
   ResetOfNotifyROS:R     "Notity_for_Rotor_over_speed";
         JU    Brake_Failure;


   //BRAKE FAILURE ALARM
   Brake_Failure:A     "Alarm_reset";
         FP    #os11;
         JC    ResetOfAlaramBF;
         CLR;
         A     "Notify_reset";
         FP    #os12;
         JC    ResetOfNotifyBF;
         CLR;
         L     "rotor_rpm";
         L     0;
         >I;
         L     "Brake_Out_HOA";
         JC    TIMERFORBF;
         JU    E_STOP;
   TIMERFORBF:CALL  "Convert_time"
         ( iv1   := "BrakeFailureSP",
           time1 := #TI_6
         );
         CALL  TON , "IEC_Timer_0_DB_24"
         ( IN := true,
           PT := #TI_6,
           Q  := #BF_AT,
           ET := #T6
         );
         A     #BF_AT;
         JC    SetOfAlarmBF;
         JU    E_STOP;

   SetOfAlarmBF:SET;
         S     "Alarm_for_Brake_failure";
         S     "Notity_for_Brake_failure";
         JU    E_STOP;
   ResetOfAlaramBF:R     "Alarm_for_Brake_failure";
         R     "Notity_for_Brake_failure";
         CALL  RESET_TIMER
         ( "TIMER" := "IEC_Timer_0_DB_24"
         );
         JU    E_STOP;
   ResetOfNotifyBF:R     "Notity_for_Brake_failure";
         JU    E_STOP;


   // E_STOP ALARM
   E_STOP:A     "Alarm_reset";
         FP    #os14;
         JC    ResetOfAlaramES;
         CLR;
         A     "Notify_reset";
         FP    #os15;
         JC    ResetOfNotifyES;
         CLR;
         A     "E_Stop";
         JC    SetOfAlarmES;
         JU    AlarmCtrl;

   SetOfAlarmES:SET;
         S     "Alarm_for_E_Stop";
         S     "Notity_for_E_Stop";
         JU    AlarmCtrl;

   ResetOfAlaramES:R     "Alarm_for_E_Stop";
         R     "Notity_for_E_Stop";
         JU    AlarmCtrl;
   ResetOfNotifyES:R     "Notity_for_E_Stop";
         JU    AlarmCtrl;

   // Alarm Horn Ctrl
   AlarmCtrl:A     "Fault_Mode";
         FP    #os16;
         JC    AlarmCtrl_SET;
         CLR;
         A     "Alarm_reset";
         O     "Notify_reset";
         FP    #os17;
         JC    ResetAlarmCtrl;
         JU    End_of_line;

   AlarmCtrl_SET:SET;
         S     "Alarm_CTRL";
         JU    End_of_line;

   ResetAlarmCtrl:R     "Alarm_CTRL";
         JU    End_of_line;

   End_of_line:BE;
END_REGION
END_FUNCTION_BLOCK

FUNCTION_BLOCK "Modes_STL"   // FB17, STL
{ S7_Optimized_Access := 'TRUE' }
VERSION : 0.1
   VAR
      os1 : Bool;
      os2 : Bool;
   END_VAR
   VAR_TEMP
      ti1 : Time;
      WarmUpTrigger : Bool;
      tm1 : Time;
      tv1 : Int;
      tv2 : Int;
      tb1 : Bool;
      ti2 : Time;
      Stabilizetrigger : Bool;
      tm2 : Time;
      ti3 : Time;
      CooldownTrigger : Bool;
      tm3 : Time;
   END_VAR
BEGIN

REGION Network 1
   // ESTOP HANDLING
         A     "Alarm_for_E_Stop";
         O     "Alarm_for_Brake_failure";
         JC    EstopAlarm;
         JU    Reset_EStopAlarm;

   EstopAlarm:SET;
         S     "Warm_Transition";
         S     "Stabilize_Transition";
         S     "Generation_Transition";
         S     "CoolDown_Transition";

   Reset_EStopAlarm:CLR;
         R     "Warm_Transition";
         R     "Stabilize_Transition";
         R     "Generation_Transition";
         R     "CoolDown_Transition";

   JumpToMode:A     "Warm_UP_Mode";
         JC    Start_WarmUp;
         CLR;
         A     "Stabilize_mode";
         JC    StabilizeMode;
         CLR;
         A     "Generation_Mode";
         JC    GenerationMode;
         CLR;
         A     "CoolDown_Mode";
         JC    CooldownMode;
         CLR;
         A     "Idle_Mode";
         JC    IdleMode;
         JU    EndOfLine;


   // WARM UP MODE
   Start_WarmUp:SET;
         R     "Warm_Transition";
         R     "Stabilize_Transition";
         R     "Generation_Transition";
         R     "CoolDown_Transition";
         R     "StartSequenceBit";
         CLR;
         A     "Warm_UP_Mode";
         JC    WarmUpMode;
         CLR;
         A     "Stabilize_mode";
         JC    StabilizeMode;
         CLR;
         A     "Generation_Mode";
         JC    GenerationMode;
         CLR;
         A     "CoolDown_Mode";
         JC    CooldownMode;
         CLR;
         A     "Idle_Mode";
         JC    IdleMode;
         JU    EndOfLine;

   WarmUpMode:SET;
         NOT;
         R     "Brake_Out_CTRL";
         L     "Warmup_RPM";
         T     "BafflePID_SP";
         L     "rotor_rpm";
         T     "BafflePIDin";

         SET;
         S     "OilPumpVFD_CTRL";
         S     "Baffle_Ctrl";
         L     "WarmUp_VFDper";
         T     "VFDsp";

         L     "Oil_temp";
         L     "WarmUpOilTempSp";
         >I;
         JC    WarmUpMode;
         CALL  RESET_TIMER
         ( "TIMER" := "IEC_Timer_0_DB_35"
         );
         JU    StabilizeMode;

   WarmUpTime:CALL  "Convert_time"
         ( iv1   := "WarmUpOilDelaySp",
           time1 := #ti1
         );
         CALL  TON, "IEC_Timer_0_DB_35"
         ( IN := true,
           PT := #ti1,
           Q  := #WarmUpTrigger,
           ET := #tm1
         );
         A     #WarmUpTrigger;
         JC    WarmUpExit;
         CLR;
         A     "Alarm_for_Rotor_over_speed";
         O     "Alarm_for_High_temp";
         JC    WarmUpExit;
         JU    StabilizeMode;

   WarmUpExit:S     "Warm_Transition";
         CALL  RESET_TIMER
         ( "TIMER" := "IEC_Timer_0_DB_35"
         );
         JU    StabilizeMode;


   //STABILZE MODE
   StabilizeMode:SET;
         NOT;
         R     "Warm_Transition";
         L     "StabilizekWSP";
         T     "BafflePID_SP";
         L     "Current_flow";
         T     "BafflePIDin";
         L     "StabilizekWSP";
         L     5;
         +I;
         T     #tv1;
         T     "StabilizekWSP";
         L     5;
         -I;
         L     #tv2;
         L     "Current_flow";
         L     #tv1;
         <I;
         S     #tb1;
         L     "Current_flow";
         L     #tv2;
         >I;
         A     #tb1;
         JC    StabilizeMode;
         CALL  RESET_TIMER
         ( "TIMER" := "IEC_Timer_0_DB_36"
         );
         JU    GenerationMode;
   StabilizeTime:CALL  "Convert_time"
         ( iv1   := "StabilizeDealySP",
           time1 := #ti2
         );
         CALL  TON, "IEC_Timer_0_DB_36"
         ( IN := true,
           PT := #ti2,
           Q  := #Stabilizetrigger,
           ET := #tm2
         );
         A     #Stabilizetrigger;
         JC    StabilizeExit;
         CLR;
         A     "Alarm_for_Rotor_over_speed";
         O     "Alarm_for_High_temp";
         JC    StabilizeExit;
         JU    GenerationMode;

   StabilizeExit:S     "Stabilize_Transition";
         CALL  RESET_TIMER
         ( "TIMER" := "IEC_Timer_0_DB_36"
         );
         JU    GenerationMode;


   //GENERATION MODE
   GenerationMode:SET;
         NOT;
         R     "Stabilize_Transition";
         SET;
         S     "Station_Interlock_CTRL";
         A     "System_Stop_PB";
         JC    GenerationExit;
         CLR;
         A     "Alarm_for_Over_Current";
         JC    GenerationExit;
         CLR;
         A     "Alarm_for_Rotor_over_speed";
         O     "Alarm_for_High_temp";
         JC    GenerationExit;
         JU    CooldownMode;

   GenerationExit:S     "Generation_Transition";
         JU    CooldownMode;


   //COOLDOWN MODE
   CooldownMode:SET;
         NOT;
         R     "Generation_Transition";
         R     "Station_Interlock_CTRL";
         L     "CoolDown_RPM";
         T     "BafflePID_SP";
         L     "rotor_rpm";
         T     "BafflePIDin";
         L     "Oil_temp";
         L     "CoolDownOilTempSp";
         <I;
         JC    Cooldowntime;
         CALL  RESET_TIMER
         ( "TIMER" := "IEC_Timer_0_DB_37"
         );
         JU    IdleMode;

   Cooldowntime:CALL  "Convert_time"
         ( iv1   := "CoolDownlDelaySp",
           time1 := #ti3
         );
         CALL  TON, "IEC_Timer_0_DB_37"
         ( IN := true,
           PT := #ti3,
           Q  := #CooldownTrigger,
           ET := #tm3
         );
         A     #CooldownTrigger;
         JC    CooldownExit;
         JU    IdleMode;

   CooldownExit:S     "CoolDown_Transition";
         CALL  RESET_TIMER
         ( "TIMER" := "IEC_Timer_0_DB_37"
         );
         JU    IdleMode;


   //IDLE MODE
   IdleMode:SET;
         NOT;
         R     "CoolDown_Transition";
         R     "Station_Interlock_CTRL";
         S     "Brake_Out_CTRL";
         R     "Baffle_Ctrl";
         R     "OilPumpVFD_CTRL";
         CLR;
         A     "StartSequencePB";
         A     "Idle_Mode";
         A     "FULLAUTOBIT";
         FP    #os2;
         S     "StartSequenceBit";
         JU    EndOfLine;

   //FAULT MODE
   EndOfLine:A     "E_Stop";
         O     "Alarm_for_Brake_failure";
         O     "Alarm_for_High_temp";
         O     "Alarm_for_LOW_OIL";
         O     "Alarm_for_Oil_High_Flow";
         O     "Alarm_for_Over_Current";
         O     "Alarm_for_Rotor_over_speed";
         =     "Fault_Mode";
END_REGION
END_FUNCTION_BLOCK

FUNCTION_BLOCK "HOURMETER_STL"   // FB22, STL
{ S7_Optimized_Access := 'TRUE' }
VERSION : 0.1
   VAR
      Min_time_down : Bool;
      Min_countdown : Bool;
      Hour_countdown : Bool;
      Day_countdown : Bool;
      Day_count_down : Bool;
      Hr_count_down : Bool;
      reset_rto : Bool;
      min_count_reset : Bool;
      hour_count_reset : Bool;
      reset_hourmeter_trigger : Bool;
      os3 : Bool;
      os2 : Bool;
      os1 : Bool;
      os4 : Bool;
      Reset_HM_Trigger : Bool;
      accum_elapsed : Time;
   END_VAR
   VAR_TEMP
      resettime : Time;
      toooomanydays : Bool;
   END_VAR
BEGIN

REGION Network 1
         A     "Generation_Mode";
         JC    RTOtimer;
         CLR;
         A     "Reset_HM_PB";
         JC    RestHourmeter;
         JU    EndOfLine;

   RTOtimer:CALL  TONR , "IEC_Timer_0_DB_44"
         ( IN := true,
           R  := #reset_rto,
           PT := t#1m,
           Q  := #Min_time_down,
           ET := #accum_elapsed
         );

         CALL  CTU, "n"
         ( CU := #Min_countdown,
           R  := #min_count_reset,
           PV := 60,
           Q  := #Hr_count_down,
           CV := "HM_Minutes"
         );

         CALL  CTU, "IEC_Counter_0_DB_9"
         ( CU := #Hour_countdown,
           R  := #hour_count_reset,
           PV := 24,
           Q  := #Day_count_down,
           CV := "HM_Hours"
         );

         CALL  CTU, "nt"
         ( CU := #Day_countdown,
           R  := #reset_hourmeter_trigger,
           PV := 10000,
           Q  := #toooomanydays,
           CV := "HM_Days"
         );

         JU    EndOfLine;

   RestHourmeter:CALL  TON, "IEC_Timer_0_DB_45"
         ( IN := "Reset_HM_PB",
           PT := T#10s,
           Q  := #Reset_HM_Trigger,
           ET := #resettime
         );

   EndOfLine:CLR;
         A     #Reset_HM_Trigger;
         O     #Min_countdown;
         =     #reset_rto;
         CLR;
         A     #Reset_HM_Trigger;
         O     #Hour_countdown;
         =     #min_count_reset;
         CLR;
         A     #Reset_HM_Trigger;
         O     #Day_countdown;
         =     #hour_count_reset;
         CLR;
END_REGION
END_FUNCTION_BLOCK

(* ===== HMI "HMI_RT_1" =====
system functions are stored by id; their names below are inferred from use
connection "1500": ETHERNET, S7_1500_OMS

HMI tags "Default tag table"
   "StartSequencePB" : Bool = PLC StartSequencePB AT %M43.7, 1 s
   "System_Stop_PB" : Bool = PLC System_Stop_PB AT %M48.7, 1 s
   "Alarm_for_E_Stop" : Bool = PLC Alarm_for_E_Stop AT %M56.0, 1 s
   "Alarm_for_Brake_failure" : Bool = PLC Alarm_for_Brake_failure AT %M55.7, 1 s
   "Alarm_for_High_temp" : Bool = PLC Alarm_for_High_temp AT %M29.7, 1 s
   "Alarm_for_LOW_OIL" : Bool = PLC Alarm_for_LOW_OIL AT %M30.0, 1 s
   "Alarm_for_Oil_High_Flow" : Bool = PLC Alarm_for_Oil_High_Flow AT %M30.1, 1 s
   "Alarm_for_Over_Current" : Bool = PLC Alarm_for_Over_Current AT %M30.2, 1 s
   "Alarm_for_Rotor_over_speed" : Bool = PLC Alarm_for_Rotor_over_speed AT %M30.3, 1 s
   "Alarm_HAND_PB" : Bool = PLC Alarm_HAND_PB AT %M28.5, 1 s
   "Alarm_HOA" : Int = PLC Alarm_HOA AT %MW34, 1 s
   "Alarm_OFF_PB" : Bool = PLC Alarm_OFF_PB AT %M28.4, 1 s
   "Alarm_reset" : Bool = PLC Alarm_reset AT %M29.6, 1 s
   "Baffle_Out" : Int = PLC Baffle_Out AT %MW18, 1 s
   "Baffle_AUTO_PB" : Bool = PLC Baffle_AUTO_PB AT %M81.2, 1 s
   "Baffle_HAND_PB" : Bool = PLC Baffle_HAND_PB AT %M81.0, 1 s
   "Baffle_HOA" : Int = PLC Baffle_HOA AT %MW94, 1 s
   "Baffle_Manual" : Bool = PLC Baffle_Manual AT %M96.0, 1 s
   "Baffle_OFF_PB" : Bool = PLC Baffle_OFF_PB AT %M81.1, 1 s
   "Brake_AUTO_PB" : Bool = PLC Brake_AUTO_PB AT %M28.3, 1 s
   "Brake_HAND_PB" : Bool = PLC Brake_HAND_PB AT %M28.2, 1 s
   "Brake_OFF_PB" : Bool = PLC Brake_OFF_PB AT %M28.1, 1 s
   "Brake_Out" : Bool = PLC Brake_Out AT %M0.0, 1 s
   "Brake_Out_CTRL" : Bool = PLC Brake_Out_CTRL AT %M29.3, 1 s
   "Brake_Out_HOA" : Int = PLC Brake_Out_HOA AT %MW32, 1 s
   "Station_interlock_HAND_PB" : Bool = PLC Station_interlock_HAND_PB AT %M29.0, 1 s
   "Station_Interlock_HOA" : Int = PLC Station_Interlock_HOA AT %MW36, 1 s
   "Station_interlock_OFF_PB" : Bool = PLC Station_interlock_OFF_PB AT %M28.7, 1 s
   "Station_interlock_AUTO_PB" : Bool = PLC Station_interlock_AUTO_PB AT %M29.1, 1 s
   "Station_interlock" : Bool = PLC Station_interlock AT %M1.3, 1 s
   "VFD_HOA" : Int = PLC VFD_HOA AT %MW98, 1 s
   "VFDHOA_AUTO_PB" : Bool = PLC VFDHOA_AUTO_PB AT %M96.1, 1 s
   "VFDHOA_HAND_PB" : Bool = PLC VFDHOA_HAND_PB AT %M96.3, 1 s
   "VFDHOA_OFF_PB" : Bool = PLC VFDHOA_OFF_PB AT %M96.2, 1 s
   "Notify_reset" : Bool = PLC Notify_reset AT %M42.1, 1 s
   "Fault_Mode" : Bool = PLC Fault_Mode AT %M80.4, 1 s
   "HighOilTempDelaySP" : Int = PLC HighOilTempDelaySP AT %MW64, 1 s
   "HM_Days" : Int = PLC HM_Days AT %MW108, 1 s
   "HM_Hours" : Int = PLC HM_Hours AT %MW106, 1 s
   "HM_Minutes" : Int = PLC HM_Minutes AT %MW30, 1 s
   "ModeInt" : Int = PLC ModeInt AT %MW110, 1 s
   "OverCurrenDelaytSP" : Int = PLC OverCurrenDelaytSP AT %MW44, 1 s
   "OilHighFlowSP" : Int = PLC OilHighFlowSP AT %MW58, 1 s
   "OilLowFlowDelaySP" : Int = PLC OilLowFlowDelaySP AT %MW38, 1 s
   "RotorOverSpeedSP" : Int = PLC RotorOverSpeedSP AT %MW54, 1 s
   "WarmUpOilTemp" : Int = PLC WarmUpOilTempSp AT %MW74, 1 s
   "CoolDownlDelaySp" : Int = PLC CoolDownlDelaySp AT %MW84, 1 s
   "CoolDownOilTemp" : Int = PLC CoolDownOilTempSp AT %MW86, 1 s
   "StabilizeDealySP" : Int = PLC StabilizeDealySP AT %MW78, 1 s
   "Alarm_horn_Q" : Bool = PLC Alarm_horn_Q AT %M1.4, 1 s
   "ManualBaffle_SP" : Real = PLC ManualBaffle_SP AT %MD90, 1 s
   "ManualVFD_SP" : Real = PLC ManualVFD_SP AT %MD100, 1 s
   "Alarm_HighOilTemp_int" : Int = PLC Alarm_HighOilTemp_int AT %MW112, 1 s
   "Alarm_LowOilFlow_int" : Int = PLC Alarm_LowOilFlow_int AT %MW114, 1 s
   "Alarm_HighOilFlow_int" : Int = PLC Alarm_HighOilFlow_int AT %MW116, 1 s
   "Alarm_OverCurrent_int" : Int = PLC Alarm_OverCurrent_int AT %MW118, 1 s
   "Alarm_RotorOverSpeed_int" : Int = PLC Alarm_RotorOverSpeed_int AT %MW120, 1 s
   "Alarm_BrakeFailure_int" : Int = PLC Alarm_BrakeFailure_int AT %MW122, 1 s
   "Alarm_EStop_int" : Int = PLC Alarm_EStop_int AT %MW124, 1 s
   "ProgramLanguage" : Int = PLC Program_lang AT %MW12, 1 s
   "LADpb" : Bool = PLC PB_LAD AT %M0.4, 1 s
   "FBDpb" : Bool = PLC PB_FBD AT %M0.5, 1 s
   "SCLpb" : Bool = PLC PB_SCL AT %M0.6, 1 s
   "STLpb" : Bool = PLC PB_STL AT %M0.7, 1 s
   "Current" : Int = PLC Current_flow AT %MW26, 1 s
   "Oil Flow" : Int = PLC Oil_flow AT %MW22, 1 s
   "Oil temp" : Int = PLC Oil_temp AT %MW24, 1 s
   "BrakeFailuredelay" : Int = PLC BrakeFailureSP AT %MW60, 1 s
   "Rpm sp" : Int = PLC Rotor_Over_SpeedSp AT %MW56, 1 s
   "OverSpeedSP" : Int = PLC RotorOverSpeedSP AT %MW54, 1 s
   "Warmup delay" : Int = PLC WarmUpOilDelaySp AT %MW72, 1 s
   "AlarmAuto_Pb" : Bool = PLC Alarm_AUTO_PB AT %M28.6, 1 s
   "RPM" : Int = PLC rotor_rpm AT %MW20, 1 s
   "OilPct" : Int = PLC Oil_pump_vfd_per AT %MW14, 1 s
   "baffle" : Int = PLC Baffle_per AT %MW16, 1 s
   "brakeEN" : Bool = PLC Brake_Out AT %M0.0, 1 s
   "InterlockEN" : Bool = PLC Station_interlock AT %M1.3, 1 s
   "HM reset" : Bool = PLC Reset_HM_PB AT %M49.0, 1 s
   "currentdealy" : Int = PLC OverCurrenDelaytSP AT %MW44, 1 s
   "high oil temp sp" : Int = PLC High_Oil_TempSp AT %MW52, 1 s
   "low oil flow sp" : Int = PLC Oil_lowSp AT %MW40, 1 s
   "curent sp" : Int = PLC Over_currentSp AT %MW46, 1 s
   "high oil flow sp" : Int = PLC Oil_highSp AT %MW62, 1 s

discrete alarms
   1: 'EStop Activated', class Errors, trigger "Alarm_EStop_int" bit 0
   2: 'Low Oil Flow Alert', class Errors, trigger "Alarm_LowOilFlow_int" bit 0
   3: 'Over Current Alert', class Errors, trigger "Alarm_OverCurrent_int" bit 0
   4: 'High Oil Temperature Alert', class Errors, trigger "Alarm_HighOilTemp_int" bit 0
   5: 'Over Speed RPM Alert', class Errors, trigger "Alarm_RotorOverSpeed_int" bit 0
   6: 'High Oil Flow Alert', class Errors, trigger "Alarm_HighOilFlow_int" bit 0
   7: 'Brake Failure Alert', class Errors, trigger "Alarm_BrakeFailure_int" bit 0

screen "Status" 1024x768
   Button "Button_1" at 42,676 size 170x70; TextOff 'Main'
      on Click: ActivateScreen("Status", 0)
   Button "Button_2" at 224,676 size 170x70; TextOff 'Overview'
      on Click: ActivateScreen("OverView", 0)
   Button "Button_3" at 404,676 size 170x70; TextOff 'Alarm'
      on Click: ActivateScreen("Alarms", 0)
   Button "Button_4" at 586,676 size 170x70; TextOff 'Config'
      on Click: ActivateScreen("Config", 0)
   TextField "Text field_3" at 12,5 size 276x61; Text 'System Status'
   TextField "Text field_4" at 605,185 size 247x62; Text 'Idle Mode'
      Visibility <- "ModeInt"
   TextField "Text field_5" at 548,185 size 361x62; Text 'WarmUp Mode'
      Visibility <- "ModeInt"
   TextField "Text field_6" at 551,185 size 356x62; Text 'Stabilize Mode'
      Visibility <- "ModeInt"
   TextField "Text field_7" at 508,185 size 442x62; Text 'Gerneration Mode'
      Visibility <- "ModeInt"
   TextField "Text field_8" at 533,185 size 391x62; Text 'Cooldown Mode'
      Visibility <- "ModeInt"
   Button "Button_5" at 624,549 size 79x62; TextOff 'LAD'
      on Press: SetBit("LADpb")
      on Release: ResetBit("LADpb")
   Button "Button_6" at 710,549 size 79x62; TextOff 'FBD'
      on Press: SetBit("FBDpb")
      on Release: ResetBit("FBDpb")
   Button "Button_7" at 796,549 size 79x62; TextOff 'SCL'
      on Press: SetBit("SCLpb")
      on Release: ResetBit("SCLpb")
   Button "Button_8" at 882,549 size 79x62; TextOff 'STL'
      on Press: SetBit("STLpb")
      on Release: ResetBit("STLpb")
   TextField "Text field_9" at 686,475 size 209x43; Text 'Ladder Logic'
      Visibility <- "ProgramLanguage"
   TextField "Text field_10" at 670,475 size 241x43; Text 'Function Block'
      Visibility <- "ProgramLanguage"
   TextField "Text field_11" at 639,475 size 302x43; Text 'Structured Control'
      Visibility <- "ProgramLanguage"
   TextField "Text field_12" at 671,475 size 238x43; Text 'Statement List'
      Visibility <- "ProgramLanguage"
   Button "Button_9" at 37,510 size 211x101; TextOff 'Start System'
      on Press: SetBit("StartSequencePB")
      on Release: ResetBit("StartSequencePB")
   Button "Button_10" at 281,510 size 211x101; TextOff 'Stop System'
      on Press: SetBit("System_Stop_PB")
      on Release: ResetBit("System_Stop_PB")
   TextField "Text field_18" at 593,83 size 239x81; Text 'MODES'
   Button "Button_11" at 857,353 size 109x43; TextOff 'Exit...'
      on Click: ActivateScreen("Config", 0)
      on Activate: StopRuntime(0)
   Group "Group_1" at 807,660 size 156x86
   Group "Group" at 806,660 size 158x86
   TextField "Text field_17" at 198,379 size 163x47; Text 'OFFLINE'
      Visibility <- "Station_interlock"
   IOField "I/O field_1" at 181,307 size 138x57; FormatPattern s99999
      ProcessValue <- "Current"
   TextField "Text field_13" at 47,312 size 128x46; Text 'Current :'
   TextField "Text field_14" at 330,314 size 49x46; Text 'kW'
   TextField "Text field_15" at 47,381 size 136x46; Text 'Interlock:'
   TextField "Text field_16" at 188,379 size 183x47; Text 'ENGAGED'
      Visibility <- "Station_interlock"
   Ellipse "Ellipse_2" at 807,660 size 156x86
      Visibility <- "Fault_Mode"
   TextField "Text field_2" at 851,676 size 70x47; Text 'OK!'
      Visibility <- "Fault_Mode"
   Ellipse "Ellipse_1" at 806,660 size 158x86
      Visibility <- "Fault_Mode"
   TextField "Text field_1" at 819,676 size 134x47; Text 'ALARM'
      Visibility <- "Fault_Mode"

screen "Alarms" 1024x768
   TextField "Text field_3" at 12,5 size 368x61; Text 'Alarm Management'
   Button "Button_1" at 42,676 size 170x70; TextOff 'Main'
      on Click: ActivateScreen("Status", 0)
   Button "Button_2" at 224,676 size 170x70; TextOff 'Overview'
      on Click: ActivateScreen("OverView", 0)
   Button "Button_3" at 404,676 size 170x70; TextOff 'Alarm'
      on Click: ActivateScreen("Alarms", 0)
   Button "Button_4" at 586,676 size 170x70; TextOff 'Config'
      on Click: ActivateScreen("Config", 0)
   AlarmView "Alarm view_1" at 25,88 size 956x194
   Group "Group_2" at 212,482 size 503x175
   Group "Group_7" at 885,319 size 126x126
   Group "Group_8" at 737,318 size 126x126
   Group "Group_9" at 589,317 size 126x126
   Group "Group_10" at 441,316 size 126x126
   Group "Group_11" at 293,315 size 126x126
   TextField "Text field_20" at 604,159 size 59x32; Text 'High'
   Group "Group_12" at 145,314 size 126x126
   Group "Group_13" at 10,317 size 126x126
   Group "Group_14" at 0,304 size 1022x154
   Group "Group_1" at 807,660 size 156x86
   Group "Group" at 806,660 size 158x86
   Circle "Circle_2" at 885,319 size 126x126
      Visibility <- "Alarm_for_LOW_OIL"
   TextField "Text field_5" at 899,365 size 101x32; Text 'Low OIL'
      Visibility <- "Alarm_for_LOW_OIL"
   Button "Button_5" at 233,566 size 216x75; TextOff 'Silence'
      on Press: SetBit("Notify_reset")
      on Release: ResetBit("Notify_reset")
   Button "Button_6" at 476,565 size 216x75; TextOff 'Alarm Reset'
      on Press: SetBit("Alarm_reset")
      on Release: ResetBit("Alarm_reset")
   TextField "Text field_6" at 360,488 size 215x46; Text 'Alarm Controls'
   Circle "Circle_1" at 737,318 size 126x126
      Visibility <- "Alarm_for_Oil_High_Flow"
   TextField "Text field_4" at 747,364 size 108x32; Text 'High OIL'
      Visibility <- "Alarm_for_Oil_High_Flow"
   Circle "Circle_3" at 589,317 size 126x126
      Visibility <- "Alarm_for_High_temp"
   Group "Group_3" at 613,347 size 69x60
   TextField "Text field_7" at 614,347 size 59x32; Text 'High'
      Visibility <- "Alarm_for_High_temp"
   TextField "Text field_14" at 613,375 size 69x32; Text 'Temp'
      Visibility <- "Alarm_for_High_temp"
   Circle "Circle_4" at 441,316 size 126x126
      Visibility <- "Alarm_for_Brake_failure"
   Group "Group_4" at 461,349 size 85x61
   TextField "Text field_8" at 461,349 size 73x32; Text 'Brake'
      Visibility <- "Alarm_for_Brake_failure"
   TextField "Text field_12" at 461,378 size 85x32; Text 'Failure'
      Visibility <- "Alarm_for_Brake_failure"
   Circle "Circle_5" at 293,315 size 126x126
      Visibility <- "Alarm_for_Over_Current"
   Group "Group_5" at 310,348 size 94x59
   TextField "Text field_9" at 312,348 size 60x32; Text 'Over'
      Visibility <- "Alarm_for_Over_Current"
   TextField "Text field_13" at 310,375 size 94x32; Text 'Current'
      Visibility <- "Alarm_for_Over_Current"
   Circle "Circle_6" at 145,314 size 126x126
      Visibility <- "Alarm_for_Rotor_over_speed"
   Group "Group_6" at 167,337 size 78x81
   TextField "Text field_10" at 167,337 size 70x32; Text 'Rotor'
      Visibility <- "Alarm_for_Rotor_over_speed"
   TextField "Text field_16" at 169,386 size 76x32; Text 'Speed'
      Visibility <- "Alarm_for_Rotor_over_speed"
   TextField "Text field_15" at 167,361 size 60x32; Text 'Over'
      Visibility <- "Alarm_for_Rotor_over_speed"
   Circle "Circle_7" at 10,317 size 126x126
      Visibility <- "Alarm_for_E_Stop"
   TextField "Text field_11" at 34,363 size 72x32; Text 'EStop'
      Visibility <- "Alarm_for_E_Stop"
   Rectangle "Rectangle_2" at 0,304 size 1022x154
      Visibility <- "Fault_Mode"
   TextField "Text field_17" at 151,332 size 673x91; Text '<<NO ALARMS>>'
      Visibility <- "Fault_Mode"
   Ellipse "Ellipse_2" at 807,660 size 156x86
      Visibility <- "Fault_Mode"
   TextField "Text field_2" at 851,676 size 70x47; Text 'OK!'
      Visibility <- "Fault_Mode"
   Ellipse "Ellipse_1" at 806,660 size 158x86
      Visibility <- "Fault_Mode"
   TextField "Text field_1" at 819,676 size 134x47; Text 'ALARM'
      Visibility <- "Fault_Mode"

screen "OverView" 1024x768
   Ellipse "Ellipse_2" at 807,660 size 156x86
      Visibility <- "Fault_Mode"
   TextField "Text field_2" at 851,676 size 70x47; Text 'OK!'
      Visibility <- "Fault_Mode"
   Ellipse "Ellipse_1" at 806,660 size 158x86
      Visibility <- "Fault_Mode"
   TextField "Text field_1" at 819,676 size 134x47; Text 'ALARM'
      Visibility <- "Fault_Mode"
   GraphicView "Graphic view_2" at 3,61 size 982x593; Picture "Graphic_1"
   TextField "Text field_3" at 12,5 size 332x61; Text 'System Overview'
   Group "Group_1" at 807,660 size 156x86
   Button "Button_1" at 42,676 size 170x70; TextOff 'Main'
      on Click: ActivateScreen("Status", 0)
   Button "Button_2" at 224,676 size 170x70; TextOff 'Overview'
      on Click: ActivateScreen("OverView", 0)
   Button "Button_3" at 404,676 size 170x70; TextOff 'Alarm'
      on Click: ActivateScreen("Alarms", 0)
   Button "Button_4" at 586,676 size 170x70; TextOff 'Config'
      on Click: ActivateScreen("Config", 0)
   Group "Group" at 806,660 size 158x86
   IOField "I/O field_1" at 25,603 size 98x37; FormatPattern s99999
      ProcessValue <- "baffle"
   TextField "Text field_4" at 25,569 size 111x36; Text 'Baffle %'
   IOField "I/O field_2" at 472,598 size 98x37; FormatPattern s99999
      ProcessValue <- "RPM"
   TextField "Text field_5" at 492,564 size 62x36; Text 'RPM'
   IOField "I/O field_3" at 556,219 size 98x37; FormatPattern s99999
      ProcessValue <- "OilPct"
   TextField "Text field_6" at 446,60 size 117x36; Text 'Oil Temp'
   TextField "Text field_7" at 811,577 size 15x22; Text 'Text'
   Group "Group_2" at 706,19 size 286x44
   Group "Group_3" at 706,19 size 286x44
   Group "Group_4" at 167,592 size 286x44
   Group "Group_5" at 167,592 size 286x44
   Group "Group_6" at 150,232 size 254x43
   TextField "Text field_12" at 819,592 size 166x43; Text 'Idle Mode'
      Visibility <- "ModeInt"
   TextField "Text field_13" at 762,592 size 243x43; Text 'WarmUp Mode'
      Visibility <- "ModeInt"
   TextField "Text field_14" at 765,592 size 240x43; Text 'Stabilize Mode'
      Visibility <- "ModeInt"
   TextField "Text field_15" at 722,592 size 294x43; Text 'Gerneration Mode'
      Visibility <- "ModeInt"
   TextField "Text field_16" at 747,592 size 261x43; Text 'Cooldown Mode'
      Visibility <- "ModeInt"
   IOField "I/O field_4" at 907,142 size 98x37; FormatPattern s99999
      ProcessValue <- "Current"
   TextField "Text field_18" at 904,106 size 99x36; Text 'Current'
   IOField "I/O field_5" at 455,94 size 98x37; FormatPattern s99999
      ProcessValue <- "Oil temp"
   Rectangle "Rectangle_1" at 167,592 size 286x44
      Visibility <- "brakeEN"
   TextField "Text field_8" at 195,596 size 232x36; Text 'Brake DisEngaged'
      Visibility <- "brakeEN"
   Rectangle "Rectangle_2" at 167,592 size 286x44
      Visibility <- "brakeEN"
   TextField "Text field_9" at 213,596 size 192x36; Text 'Brake Engaged'
      Visibility <- "brakeEN"
   Rectangle "Rectangle_3" at 706,19 size 286x44
      Visibility <- "InterlockEN"
   TextField "Text field_10" at 735,23 size 233x36; Text 'Interlock Engaged'
      Visibility <- "InterlockEN"
   Rectangle "Rectangle_4" at 706,19 size 286x44
      Visibility <- "InterlockEN"
   TextField "Text field_11" at 712,23 size 273x36; Text 'Interlock DisEngaged'
      Visibility <- "InterlockEN"
   Rectangle "Rectangle_5" at 150,232 size 254x43
      Visibility <- "Fault_Mode"
   TextField "Text field_17" at 166,235 size 222x32; Text '<<NO ALARMS>>'

screen "Config" 1024x768
   TextField "Text field_3" at 12,5 size 262x61; Text 'Configuration'
   Button "Button_1" at 42,676 size 170x70; TextOff 'Main'
      on Click: ActivateScreen("Status", 0)
   Button "Button_2" at 224,676 size 170x70; TextOff 'Overview'
      on Click: ActivateScreen("OverView", 0)
   Button "Button_3" at 404,676 size 170x70; TextOff 'Alarm'
      on Click: ActivateScreen("Alarms", 0)
   Button "Button_4" at 586,676 size 170x70; TextOff 'Config'
      on Click: ActivateScreen("Config", 0)
   Group "Group_9" at 397,418 size 169x203
   Group "Group_1" at 807,660 size 156x86
   Group "Group" at 806,660 size 158x86
   Group "Group_2" at 9,90 size 321x526
   Group "Group_3" at 345,88 size 302x315
   Group "Group_4" at 664,89 size 344x540
   TextField "Text field_4" at 18,93 size 172x41; Text 'Alarm Values'
   TextField "Text field_5" at 18,138 size 210x37; Text 'Brake Failure Delay'
   IOField "I/O field_9" at 232,137 size 76x38; FormatPattern 99999
      ProcessValue <- "BrakeFailuredelay"
   TextField "Text field_6" at 18,181 size 123x37; Text 'Rotor RPM'
   IOField "I/O field_1" at 232,180 size 76x38; FormatPattern s99999
      ProcessValue <- "RPM"
   TextField "Text field_7" at 18,224 size 171x37; Text 'Rotor RPM (sp)'
   IOField "I/O field_2" at 232,223 size 76x38; FormatPattern s99999
      ProcessValue <- "Rpm sp"
   TextField "Text field_8" at 18,267 size 205x37; Text 'High Oil Temp (sp)'
   IOField "I/O field_3" at 232,266 size 76x38; FormatPattern s99999
      ProcessValue <- "high oil temp sp"
   TextField "Text field_9" at 18,310 size 186x37; Text 'Oil Temp Degree'
   IOField "I/O field_4" at 232,309 size 76x38; FormatPattern s99999
      ProcessValue <- "Oil temp"
   TextField "Text field_10" at 18,353 size 187x37; Text 'Low Oil Flow (sp)'
   IOField "I/O field_5" at 232,352 size 76x38; FormatPattern s99999
      ProcessValue <- "low oil flow sp"
   TextField "Text field_11" at 18,396 size 167x37; Text 'Oil Flow (GPM)'
   IOField "I/O field_6" at 232,395 size 76x38; FormatPattern s99999
      ProcessValue <- "Oil Flow"
   TextField "Text field_12" at 18,439 size 193x37; Text 'High Oil Flow (sp)'
   IOField "I/O field_7" at 232,438 size 76x38; FormatPattern s99999
      ProcessValue <- "high oil flow sp"
   TextField "Text field_13" at 18,482 size 167x37; Text 'Oil Flow (GPM)'
   IOField "I/O field_8" at 232,481 size 76x38; FormatPattern s99999
      ProcessValue <- "Oil Flow"
   TextField "Text field_33" at 18,526 size 141x37; Text 'Current (kW)'
   IOField "I/O field_20" at 232,525 size 76x38; FormatPattern s99999
      ProcessValue <- "Current"
   TextField "Text field_34" at 18,569 size 132x37; Text 'Current (sp)'
   IOField "I/O field_21" at 232,568 size 76x38; FormatPattern s99999
      ProcessValue <- "curent sp"
   TextField "Text field_14" at 353,91 size 202x41; Text 'Process Values'
   TextField "Text field_15" at 353,136 size 162x37; Text 'Warmup Temp'
   IOField "I/O field_10" at 534,135 size 90x38; FormatPattern 99999
      ProcessValue <- "WarmUpOilTemp"
   TextField "Text field_16" at 353,179 size 159x37; Text 'Warmup Delay'
   IOField "I/O field_11" at 534,178 size 90x38; FormatPattern s99999
      ProcessValue <- "Warmup delay"
   TextField "Text field_17" at 353,222 size 141x37; Text 'Current (kW)'
   IOField "I/O field_12" at 534,221 size 90x38; FormatPattern s99999
      ProcessValue <- "Current"
   TextField "Text field_18" at 353,265 size 158x37; Text 'Stabilize Delay'
   IOField "I/O field_13" at 534,264 size 90x38; FormatPattern s99999
      ProcessValue <- "StabilizeDealySP"
   TextField "Text field_19" at 353,308 size 177x37; Text 'Cooldown Temp'
   IOField "I/O field_14" at 534,307 size 90x38; FormatPattern s99999
      ProcessValue <- "CoolDownOilTemp"
   TextField "Text field_20" at 353,351 size 174x37; Text 'Cooldown Delay'
   IOField "I/O field_15" at 534,350 size 90x38; FormatPattern s99999
      ProcessValue <- "CoolDownlDelaySp"
   Rectangle "Rectangle_7" at 674,233 size 324x80
      Visibility <- "Brake_Out_HOA"
   Rectangle "Rectangle_8" at 674,233 size 324x80
      Visibility <- "Brake_Out_HOA"
   Rectangle "Rectangle_9" at 674,233 size 324x80
      Visibility <- "Brake_Out_HOA"
   Rectangle "Rectangle_4" at 673,145 size 324x80
      Visibility <- "Alarm_HOA"
   Rectangle "Rectangle_5" at 673,145 size 324x80
      Visibility <- "Alarm_HOA"
   Rectangle "Rectangle_6" at 673,145 size 324x80
      Visibility <- "Alarm_HOA"
   TextField "Text field_21" at 674,91 size 178x41; Text 'HOA Controls'
   Rectangle "Rectangle_10" at 674,517 size 324x100
      Visibility <- "VFD_HOA"
   Rectangle "Rectangle_11" at 674,517 size 324x100
      Visibility <- "VFD_HOA"
   Rectangle "Rectangle_12" at 674,517 size 324x100
      Visibility <- "VFD_HOA"
   Rectangle "Rectangle_13" at 674,321 size 324x80
      Visibility <- "Station_Interlock_HOA"
   Rectangle "Rectangle_14" at 674,321 size 324x80
      Visibility <- "Station_Interlock_HOA"
   Rectangle "Rectangle_15" at 674,321 size 324x80
      Visibility <- "Station_Interlock_HOA"
   Rectangle "Rectangle_16" at 674,408 size 324x100
      Visibility <- "Baffle_HOA"
   Rectangle "Rectangle_17" at 674,408 size 324x100
      Visibility <- "Baffle_HOA"
   Rectangle "Rectangle_18" at 674,408 size 324x100
      Visibility <- "Baffle_HOA"
   TextField "Text field_24" at 682,323 size 126x34; Text 'InterLock'
   Button "Button_11" at 683,361 size 96x39; TextOff 'Hand'
      on Press: SetBit("Station_interlock_HAND_PB")
      on Release: ResetBit("Station_interlock_HAND_PB")
   Button "Button_12" at 788,360 size 96x39; TextOff 'OFF'
      on Release: ResetBit("Station_interlock_OFF_PB")
      on Press: SetBit("Station_interlock_OFF_PB")
   Button "Button_13" at 893,360 size 96x39; TextOff 'AUTO'
      on Press: SetBit("Station_interlock_AUTO_PB")
      on Release: ResetBit("Station_interlock_AUTO_PB")
   IOField "I/O field_16" at 899,538 size 99x44; FormatPattern s99999
      ProcessValue <- "ManualVFD_SP"
   TextField "Text field_28" at 908,516 size 82x22; Text 'Manual Sp'
   TextField "Text field_27" at 687,523 size 177x34; Text 'Oil Pump VFD'
   Button "Button_18" at 788,584 size 96x32; TextOff 'OFF'
      on Release: ResetBit("VFDHOA_HAND_PB")
      on Press: SetBit("VFDHOA_HAND_PB")
   Button "Button_19" at 893,584 size 96x32; TextOff 'AUTO'
      on Press: SetBit("VFDHOA_AUTO_PB")
      on Release: ResetBit("VFDHOA_AUTO_PB")
   Button "Button_17" at 683,585 size 96x32; TextOff 'Hand'
      on Press: SetBit("VFDHOA_HAND_PB")
      on Release: ResetBit("VFDHOA_HAND_PB")
   TextField "Text field_23" at 681,236 size 78x34; Text 'Brake'
   Button "Button_9" at 683,273 size 96x39; TextOff 'Hand'
      on Press: SetBit("Brake_HAND_PB")
      on Release: ResetBit("Brake_HAND_PB")
   Button "Button_10" at 788,272 size 96x39; TextOff 'OFF'
      on Release: ResetBit("Brake_OFF_PB")
      on Press: SetBit("Brake_OFF_PB")
   Button "Button_8" at 893,272 size 96x39; TextOff 'AUTO'
      on Press: SetBit("Brake_AUTO_PB")
      on Release: ResetBit("Brake_AUTO_PB")
   Button "Button_5" at 681,186 size 96x40; TextOff 'Hand'
      on Press: SetBit("Alarm_HAND_PB")
      on Release: ResetBit("Alarm_HAND_PB")
   TextField "Text field_22" at 681,147 size 148x34; Text 'Alarm Horn'
   Button "Button_6" at 786,185 size 96x40; TextOff 'OFF'
      on Release: ResetBit("Alarm_OFF_PB")
      on Press: SetBit("Alarm_OFF_PB")
   Button "Button_7" at 891,185 size 96x40; TextOff 'AUTO'
      on Press: SetBit("AlarmAuto_Pb")
      on Release: ResetBit("AlarmAuto_Pb")
   IOField "I/O field_23" at 900,429 size 99x44; FormatPattern s999999999.999
      ProcessValue <- "ManualBaffle_SP"
   TextField "Text field_26" at 909,407 size 82x22; Text 'Manual Sp'
   Button "Button_16" at 897,476 size 96x32; TextOff 'AUTO'
      on Press: SetBit("Baffle_AUTO_PB")
      on Release: ResetBit("Baffle_AUTO_PB")
   Button "Button_15" at 792,476 size 96x32; TextOff 'OFF'
      on Release: ResetBit("Baffle_OFF_PB")
      on Press: SetBit("Baffle_OFF_PB")
   Button "Button_14" at 687,477 size 96x32; TextOff 'Hand'
      on Press: SetBit("Baffle_HAND_PB")
      on Release: ResetBit("Baffle_HAND_PB")
   TextField "Text field_25" at 682,414 size 80x34; Text 'Baffle'
   IOField "I/O field_17" at 470,457 size 96x32; FormatPattern s99999
      ProcessValue <- "HM_Days"
   TextField "Text field_29" at 412,418 size 138x32; Text 'Hour Meter'
   TextField "Text field_30" at 402,457 size 57x29; Text 'Days'
   IOField "I/O field_18" at 470,499 size 96x32; FormatPattern s99999
      ProcessValue <- "HM_Hours"
   TextField "Text field_31" at 397,499 size 67x29; Text 'Hours'
   IOField "I/O field_19" at 470,541 size 96x32; FormatPattern s99999
      ProcessValue <- "HM_Minutes"
   TextField "Text field_32" at 406,541 size 54x29; Text 'Mins'
   Button "Button_20" at 433,581 size 106x40; TextOff 'HM Reset'
      on Press: SetBit("HM reset")
      on Release: ResetBit("HM reset")
   Ellipse "Ellipse_2" at 807,660 size 156x86
      Visibility <- "Fault_Mode"
   TextField "Text field_2" at 851,676 size 70x47; Text 'OK!'
      Visibility <- "Fault_Mode"
   Ellipse "Ellipse_1" at 806,660 size 158x86
      Visibility <- "Fault_Mode"
   TextField "Text field_1" at 819,676 size 134x47; Text 'ALARM'
      Visibility <- "Fault_Mode"
*)